   15328: 'Mixinghead 04: Cleaning piston: Front position not reached', class Mixing Head Warning, trigger "Mixinghead_Cpiston4_DBW_40" bit 3
   15329: 'Mixinghead 04: Cleaning piston: Rear position not reached', class Mixing Head Warning, trigger "Mixinghead_Cpiston4_DBW_40" bit 4
   15330: 'Mixinghead 04: Cleaning piston: Home position not reached', class Mixing Head Warning, trigger "Mixinghead_Cpiston4_DBW_40" bit 5
   15331: 'Mixinghead 04: Cleaning piston:', class Mixing Head Warning, trigger "Mixinghead_Cpiston4_DBW_40" bit 6
   15332: 'Mixinghead 04: Cleaning piston:', class Mixing Head Warning, trigger "Mixinghead_Cpiston4_DBW_40" bit 7
   15340: 'Mixinghead 04: Connection 01: Temperature recording: Measuring value outside measuring range', class Mixing Head Warning, trigger "Mixinghead_Temperature_MH4_Con1_DBW76" bit 8
   15341: 'Mixinghead 04: Connection 01: Temperature recording: Warning, value exceeded', class Mixing Head Warning, trigger "Mixinghead_Temperature_MH4_Con1_DBW76" bit 9
   15342: 'Mixinghead 04: Connection 01: Temperature recording: Warning, value undershot', class Mixing Head Warning, trigger "Mixinghead_Temperature_MH4_Con1_DBW76" bit 10
   15343: 'Mixinghead 04: Connection 01: Temperature recording: Fault, value exceeded', class Mixing Head Errors, trigger "Mixinghead_Temperature_MH4_Con1_DBW76" bit 11
   15344: 'Mixinghead 04: Connection 01: Temperature recording: Fault, value undershot', class Mixing Head Errors, trigger "Mixinghead_Temperature_MH4_Con1_DBW76" bit 12
   15345: 'Mixinghead 04: Connection 02: Temperature recording: Measuring value outside measuring range', class Mixing Head Warning, trigger "Mixinghead_Temperature_MH4_Con2_DBW110" bit 8
   15346: 'Mixinghead 04: Connection 02: Temperature recording: Warning, value exceeded', class Mixing Head Warning, trigger "Mixinghead_Temperature_MH4_Con2_DBW110" bit 9
   15347: 'Mixinghead 04: Connection 02: Temperature recording: Warning, value undershot', class Mixing Head Warning, trigger "Mixinghead_Temperature_MH4_Con2_DBW110" bit 10
   15348: 'Mixinghead 04: Connection 02: Temperature recording: Fault, value exceeded', class Mixing Head Errors, trigger "Mixinghead_Temperature_MH4_Con2_DBW110" bit 11
   15349: 'Mixinghead 04: Connection 02: Temperature recording: Fault, value undershot', class Mixing Head Errors, trigger "Mixinghead_Temperature_MH4_Con2_DBW110" bit 12
   15350: 'Mixinghead 04: Connection 03: Temperature recording: Measuring value outside measuring range', class Mixing Head Warning, trigger "Mixinghead_Temperature_MH4_Con3_DBW144" bit 8
   15351: 'Mixinghead 04: Connection 03: Temperature recording: Warning, value exceeded', class Mixing Head Warning, trigger "Mixinghead_Temperature_MH4_Con3_DBW144" bit 9
   15352: 'Mixinghead 04: Connection 03: Temperature recording: Warning, value undershot', class Mixing Head Warning, trigger "Mixinghead_Temperature_MH4_Con3_DBW144" bit 10
   15353: 'Mixinghead 04: Connection 03: Temperature recording: Fault, value exceeded', class Mixing Head Errors, trigger "Mixinghead_Temperature_MH4_Con3_DBW144" bit 11
   15354: 'Mixinghead 04: Connection 03: Temperature recording: Fault, value undershot', class Mixing Head Errors, trigger "Mixinghead_Temperature_MH4_Con3_DBW144" bit 12
   15355: 'Mixinghead 04: Connection 04: Temperature recording: Measuring value outside measuring range', class Mixing Head Warning, trigger "Mixinghead_Temperature_MH4_Con4_DBW178" bit 8
   15356: 'Mixinghead 04: Connection 04: Temperature recording: Warning, value exceeded', class Mixing Head Warning, trigger "Mixinghead_Temperature_MH4_Con4_DBW178" bit 9
   15357: 'Mixinghead 04: Connection 04: Temperature recording: Warning, value undershot', class Mixing Head Warning, trigger "Mixinghead_Temperature_MH4_Con4_DBW178" bit 10
   15358: 'Mixinghead 04: Connection 04: Temperature recording: Fault, value exceeded', class Mixing Head Errors, trigger "Mixinghead_Temperature_MH4_Con4_DBW178" bit 11
   15359: 'Mixinghead 04: Connection 04: Temperature recording: Fault, value undershot', class Mixing Head Errors, trigger "Mixinghead_Temperature_MH4_Con4_DBW178" bit 12
   15360: 'Mixinghead 04: Connection 05: Temperature recording: Measuring value outside measuring range', class Mixing Head Warning, trigger "Mixinghead_Temperature_MH4_Con5_DBW212" bit 8
   15361: 'Mixinghead 04: Connection 05: Temperature recording: Warning, value exceeded', class Mixing Head Warning, trigger "Mixinghead_Temperature_MH4_Con5_DBW212" bit 9
   15362: 'Mixinghead 04: Connection 05: Temperature recording: Warning, value undershot', class Mixing Head Warning, trigger "Mixinghead_Temperature_MH4_Con5_DBW212" bit 10
   15363: 'Mixinghead 04: Connection 05: Temperature recording: Fault, value exceeded', class Mixing Head Errors, trigger "Mixinghead_Temperature_MH4_Con5_DBW212" bit 11
   15364: 'Mixinghead 04: Connection 05: Temperature recording: Fault, value undershot', class Mixing Head Errors, trigger "Mixinghead_Temperature_MH4_Con5_DBW212" bit 12
   15365: 'Mixinghead 04: Connection 06: Temperature recording: Measuring value outside measuring range', class Mixing Head Warning, trigger "Mixinghead_Temperature_MH4_Con6_DBW246" bit 8
   15366: 'Mixinghead 04: Connection 06: Temperature recording: Warning, value exceeded', class Mixing Head Warning, trigger "Mixinghead_Temperature_MH4_Con6_DBW246" bit 9
   15367: 'Mixinghead 04: Connection 06: Temperature recording: Warning, value undershot', class Mixing Head Warning, trigger "Mixinghead_Temperature_MH4_Con6_DBW246" bit 10
   15368: 'Mixinghead 04: Connection 06: Temperature recording: Fault, value exceeded', class Mixing Head Errors, trigger "Mixinghead_Temperature_MH4_Con6_DBW246" bit 11
   15369: 'Mixinghead 04: Connection 06: Temperature recording: Fault, value undershot', class Mixing Head Errors, trigger "Mixinghead_Temperature_MH4_Con6_DBW246" bit 12
   15370: 'Mixinghead 04: Connection 01: Pressure recording: Measuring value outside measuring range', class Mixing Head Warning, trigger "Mixinghead_Pressure_MH4_Con1_DBW280" bit 8
   15371: 'Mixinghead 04: Connection 01: Pressure recording: Warning, value exceeded', class Mixing Head Warning, trigger "Mixinghead_Pressure_MH4_Con1_DBW280" bit 9
   15372: 'Mixinghead 04: Connection 01: Pressure recording: Warning, value undershot', class Mixing Head Warning, trigger "Mixinghead_Pressure_MH4_Con1_DBW280" bit 10
   15373: 'Mixinghead 04: Connection 01: Pressure recording: Fault, value exceeded', class Mixing Head Errors, trigger "Mixinghead_Pressure_MH4_Con1_DBW280" bit 11
   15374: 'Mixinghead 04: Connection 01: Pressure recording: Fault, value undershot', class Mixing Head Errors, trigger "Mixinghead_Pressure_MH4_Con1_DBW280" bit 12
   15375: 'Mixinghead 04: Connection 02: Pressure recording: Measuring value outside measuring range', class Mixing Head Warning, trigger "Mixinghead_Pressure_MH4_Con2_DBW314" bit 8
   15376: 'Mixinghead 04: Connection 02: Pressure recording: Warning, value exceeded', class Mixing Head Warning, trigger "Mixinghead_Pressure_MH4_Con2_DBW314" bit 9
   15377: 'Mixinghead 04: Connection 02: Pressure recording: Warning, value undershot', class Mixing Head Warning, trigger "Mixinghead_Pressure_MH4_Con2_DBW314" bit 10
   15378: 'Mixinghead 04: Connection 02: Pressure recording: Fault, value exceeded', class Mixing Head Errors, trigger "Mixinghead_Pressure_MH4_Con2_DBW314" bit 11
   15379: 'Mixinghead 04: Connection 02: Pressure recording: Fault, value undershot', class Mixing Head Errors, trigger "Mixinghead_Pressure_MH4_Con2_DBW314" bit 12
   15380: 'Mixinghead 04: Connection 03: Pressure recording: Measuring value outside measuring range', class Mixing Head Warning, trigger "Mixinghead_Pressure_MH4_Con3_DBW348" bit 8
   15381: 'Mixinghead 04: Connection 03: Pressure recording: Warning, value exceeded', class Mixing Head Warning, trigger "Mixinghead_Pressure_MH4_Con3_DBW348" bit 9
   15382: 'Mixinghead 04: Connection 03: Pressure recording: Warning, value undershot', class Mixing Head Warning, trigger "Mixinghead_Pressure_MH4_Con3_DBW348" bit 10
   15383: 'Mixinghead 04: Connection 03: Pressure recording: Fault, value exceeded', class Mixing Head Errors, trigger "Mixinghead_Pressure_MH4_Con3_DBW348" bit 11
   15384: 'Mixinghead 04: Connection 03: Pressure recording: Fault, value undershot', class Mixing Head Errors, trigger "Mixinghead_Pressure_MH4_Con3_DBW348" bit 12
   15385: 'Mixinghead 04: Connection 04: Pressure recording: Measuring value outside measuring range', class Mixing Head Warning, trigger "Mixinghead_Pressure_MH4_Con4_DBW382" bit 8
   15386: 'Mixinghead 04: Connection 04: Pressure recording: Warning, value exceeded', class Mixing Head Warning, trigger "Mixinghead_Pressure_MH4_Con4_DBW382" bit 9
   15387: 'Mixinghead 04: Connection 04: Pressure recording: Warning, value undershot', class Mixing Head Warning, trigger "Mixinghead_Pressure_MH4_Con4_DBW382" bit 10
   15388: 'Mixinghead 04: Connection 04: Pressure recording: Fault, value exceeded', class Mixing Head Errors, trigger "Mixinghead_Pressure_MH4_Con4_DBW382" bit 11
   15389: 'Mixinghead 04: Connection 04: Pressure recording: Fault, value undershot', class Mixing Head Errors, trigger "Mixinghead_Pressure_MH4_Con4_DBW382" bit 12
   15390: 'Mixinghead 04: Connection 05: Pressure recording: Measuring value outside measuring range', class Mixing Head Warning, trigger "Mixinghead_Pressure_MH4_Con5_DBW416" bit 8
   15391: 'Mixinghead 04: Connection 05: Pressure recording: Warning, value exceeded', class Mixing Head Warning, trigger "Mixinghead_Pressure_MH4_Con5_DBW416" bit 9
   15392: 'Mixinghead 04: Connection 05: Pressure recording: Warning, value undershot', class Mixing Head Warning, trigger "Mixinghead_Pressure_MH4_Con5_DBW416" bit 10
   15393: 'Mixinghead 04: Connection 05: Pressure recording: Fault, value exceeded', class Mixing Head Errors, trigger "Mixinghead_Pressure_MH4_Con5_DBW416" bit 11
   15394: 'Mixinghead 04: Connection 05: Pressure recording: Fault, value undershot', class Mixing Head Errors, trigger "Mixinghead_Pressure_MH4_Con5_DBW416" bit 12
   15395: 'Mixinghead 04: Connection 06: Pressure recording: Measuring value outside measuring range', class Mixing Head Warning, trigger "Mixinghead_Pressure_MH4_Con6_DBW450" bit 8
   15396: 'Mixinghead 04: Connection 06: Pressure recording: Warning, value exceeded', class Mixing Head Warning, trigger "Mixinghead_Pressure_MH4_Con6_DBW450" bit 9
   15397: 'Mixinghead 04: Connection 06: Pressure recording: Warning, value undershot', class Mixing Head Warning, trigger "Mixinghead_Pressure_MH4_Con6_DBW450" bit 10
   15398: 'Mixinghead 04: Connection 06: Pressure recording: Fault, value exceeded', class Mixing Head Errors, trigger "Mixinghead_Pressure_MH4_Con6_DBW450" bit 11
   15399: 'Mixinghead 04: Connection 06: Pressure recording: Fault, value undershot', class Mixing Head Errors, trigger "Mixinghead_Pressure_MH4_Con6_DBW450" bit 12
   15401: 'Mixinghead 05: Mixinghead does not open', class Mixing Head Errors, trigger "Mixinghead_MHControl5_DBW_10" bit 8
   15402: 'Mixinghead 05: Mixinghead does not close', class Mixing Head Errors, trigger "Mixinghead_MHControl5_DBW_10" bit 9
   15403: 'Mixinghead 05: Entry cancelled', class Mixing Head Warning, trigger "Mixinghead_MHControl5_DBW_10" bit 10
   15404: 'Mixinghead 05: Mixinghead open without activation', class Mixing Head Errors, trigger "Mixinghead_MHControl5_DBW_10" bit 11
   15405: 'Mixinghead 05: Mixinghead close during entry', class Mixing Head Warning, trigger "Mixinghead_MHControl5_DBW_10" bit 12
   15406: 'Mixinghead 05: Warning, shot time too short', class Mixing Head Warning, trigger "Mixinghead_MHControl5_DBW_10" bit 13
   15407: 'Mixinghead 05: Warning , shot time too long', class Mixing Head Warning, trigger "Mixinghead_MHControl5_DBW_10" bit 14
   15408: 'Mixinghead 05: Fault, shot time too short', class Mixing Head Warning, trigger "Mixinghead_MHControl5_DBW_10" bit 15
   15409: 'Mixinghead 05: Mixinghead collides when opening or closing', class Mixing Head Warning, trigger "Mixinghead_MHControl5_DBW_10" bit 0
   15410: 'Mixinghead 05: Runtime monitoring when locking mixing head', class Mixing Head Warning, trigger "Mixinghead_MHControl5_DBW_10" bit 1
   15411: 'Mixinghead 05: Runtime monitoring when unlocking mixing head', class Mixing Head Warning, trigger "Mixinghead_MHControl5_DBW_10" bit 2
   15412: 'Mixinghead 05:', class Mixing Head Warning, trigger "Mixinghead_MHControl5_DBW_10" bit 3
   15413: 'Mixinghead 05:', class Mixing Head Warning, trigger "Mixinghead_MHControl5_DBW_10" bit 4
   15414: 'Mixinghead 05:', class Mixing Head Warning, trigger "Mixinghead_MHControl5_DBW_10" bit 5
   15415: 'Mixinghead 05:', class Mixing Head Warning, trigger "Mixinghead_MHControl5_DBW_10" bit 6
   15416: 'Mixinghead 05: Component required in entry is not enabled at this mixing head', class Mixing Head Errors, trigger "Mixinghead_MHControl5_DBW_10" bit 7
   15417: 'Mixinghead 05: Cleaning piston: Moving out too slow', class Mixing Head Errors, trigger "Mixinghead_Cpiston5_DBW_42" bit 8
   15418: 'Mixinghead 05: Cleaning piston: Moving in too slow', class Mixing Head Errors, trigger "Mixinghead_Cpiston5_DBW_42" bit 9
   15419: 'Mixinghead 05: Cleaning piston: Proximity switch defect', class Mixing Head Errors, trigger "Mixinghead_Cpiston5_DBW_42" bit 10
   15420: 'Mixinghead 05: Cleaning piston: Leaves its home position in entry', class Mixing Head Errors, trigger "Mixinghead_Cpiston5_DBW_42" bit 11
   15421: 'Mixinghead 05: Cleaning piston: Not defined', class Mixing Head Warning, trigger "Mixinghead_Cpiston5_DBW_42" bit 12
   15422: 'Mixinghead 05: Cleaning piston:', class Mixing Head Warning, trigger "Mixinghead_Cpiston5_DBW_42" bit 13
   15423: 'Mixinghead 05: Cleaning piston:', class Mixing Head Warning, trigger "Mixinghead_Cpiston5_DBW_42" bit 14
   15424: 'Mixinghead 05: Cleaning piston:', class Mixing Head Warning, trigger "Mixinghead_Cpiston5_DBW_42" bit 15
   15425: 'Mixinghead 05: Cleaning piston: Controller at upper limit', class Mixing Head Warning, trigger "Mixinghead_Cpiston5_DBW_42" bit 0
   15426: 'Mixinghead 05: Cleaning piston: Controller at lower limit', class Mixing Head Warning, trigger "Mixinghead_Cpiston5_DBW_42" bit 1
   15427: 'Mixinghead 05: Cleaning piston:', class Mixing Head Warning, trigger "Mixinghead_Cpiston5_DBW_42" bit 2
   15428: 'Mixinghead 05: Cleaning piston: Front position not reached', class Mixing Head Warning, trigger "Mixinghead_Cpiston5_DBW_42" bit 3
   15429: 'Mixinghead 05: Cleaning piston: Rear position not reached', class Mixing Head Warning, trigger "Mixinghead_Cpiston5_DBW_42" bit 4
   15430: 'Mixinghead 05: Cleaning piston: Home position not reached', class Mixing Head Warning, trigger "Mixinghead_Cpiston5_DBW_42" bit 5
   15431: 'Mixinghead 05: Cleaning piston:', class Mixing Head Warning, trigger "Mixinghead_Cpiston5_DBW_42" bit 6
   15432: 'Mixinghead 05: Cleaning piston:', class Mixing Head Warning, trigger "Mixinghead_Cpiston5_DBW_42" bit 7
   15440: 'Mixinghead 05: Connection 01: Temperature recording: Measuring value outside measuring range', class Mixing Head Warning, trigger "Mixinghead_Temperature_MH5_Con1_DBW78" bit 8
   15441: 'Mixinghead 05: Connection 01: Temperature recording: Warning, value exceeded', class Mixing Head Warning, trigger "Mixinghead_Temperature_MH5_Con1_DBW78" bit 9
   15442: 'Mixinghead 05: Connection 01: Temperature recording: Warning, value undershot', class Mixing Head Warning, trigger "Mixinghead_Temperature_MH5_Con1_DBW78" bit 10
   15443: 'Mixinghead 05: Connection 01: Temperature recording: Fault, value exceeded', class Mixing Head Errors, trigger "Mixinghead_Temperature_MH5_Con1_DBW78" bit 11
   15444: 'Mixinghead 05: Connection 01: Temperature recording: Fault, value undershot', class Mixing Head Errors, trigger "Mixinghead_Temperature_MH5_Con1_DBW78" bit 12
   15445: 'Mixinghead 05: Connection 02: Temperature recording: Measuring value outside measuring range', class Mixing Head Warning, trigger "Mixinghead_Temperature_MH5_Con2_DBW112" bit 8
   15446: 'Mixinghead 05: Connection 02: Temperature recording: Warning, value exceeded', class Mixing Head Warning, trigger "Mixinghead_Temperature_MH5_Con2_DBW112" bit 9
   15447: 'Mixinghead 05: Connection 02: Temperature recording: Warning, value undershot', class Mixing Head Warning, trigger "Mixinghead_Temperature_MH5_Con2_DBW112" bit 10
   15448: 'Mixinghead 05: Connection 02: Temperature recording: Fault, value exceeded', class Mixing Head Errors, trigger "Mixinghead_Temperature_MH5_Con2_DBW112" bit 11
   15449: 'Mixinghead 05: Connection 02: Temperature recording: Fault, value undershot', class Mixing Head Errors, trigger "Mixinghead_Temperature_MH5_Con2_DBW112" bit 12
   15450: 'Mixinghead 05: Connection 03: Temperature recording: Measuring value outside measuring range', class Mixing Head Warning, trigger "Mixinghead_Temperature_MH5_Con3_DBW146" bit 8
   15451: 'Mixinghead 05: Connection 03: Temperature recording: Warning, value exceeded', class Mixing Head Warning, trigger "Mixinghead_Temperature_MH5_Con3_DBW146" bit 9
   15452: 'Mixinghead 05: Connection 03: Temperature recording: Warning, value undershot', class Mixing Head Warning, trigger "Mixinghead_Temperature_MH5_Con3_DBW146" bit 10
   15453: 'Mixinghead 05: Connection 03: Temperature recording: Fault, value exceeded', class Mixing Head Errors, trigger "Mixinghead_Temperature_MH5_Con3_DBW146" bit 11
   15454: 'Mixinghead 05: Connection 03: Temperature recording: Fault, value undershot', class Mixing Head Errors, trigger "Mixinghead_Temperature_MH5_Con3_DBW146" bit 12
   15455: 'Mixinghead 05: Connection 04: Temperature recording: Measuring value outside measuring range', class Mixing Head Warning, trigger "Mixinghead_Temperature_MH5_Con4_DBW180" bit 8
   15456: 'Mixinghead 05: Connection 04: Temperature recording: Warning, value exceeded', class Mixing Head Warning, trigger "Mixinghead_Temperature_MH5_Con4_DBW180" bit 9
   15457: 'Mixinghead 05: Connection 04: Temperature recording: Warning, value undershot', class Mixing Head Warning, trigger "Mixinghead_Temperature_MH5_Con4_DBW180" bit 10
   15458: 'Mixinghead 05: Connection 04: Temperature recording: Fault, value exceeded', class Mixing Head Errors, trigger "Mixinghead_Temperature_MH5_Con4_DBW180" bit 11
   15459: 'Mixinghead 05: Connection 04: Temperature recording: Fault, value undershot', class Mixing Head Errors, trigger "Mixinghead_Temperature_MH5_Con4_DBW180" bit 12
   15460: 'Mixinghead 05: Connection 05: Temperature recording: Measuring value outside measuring range', class Mixing Head Warning, trigger "Mixinghead_Temperature_MH5_Con5_DBW214" bit 8
   15461: 'Mixinghead 05: Connection 05: Temperature recording: Warning, value exceeded', class Mixing Head Warning, trigger "Mixinghead_Temperature_MH5_Con5_DBW214" bit 9
   15462: 'Mixinghead 05: Connection 05: Temperature recording: Warning, value undershot', class Mixing Head Warning, trigger "Mixinghead_Temperature_MH5_Con5_DBW214" bit 10
   15463: 'Mixinghead 05: Connection 05: Temperature recording: Fault, value exceeded', class Mixing Head Errors, trigger "Mixinghead_Temperature_MH5_Con5_DBW214" bit 11
   15464: 'Mixinghead 05: Connection 05: Temperature recording: Fault, value undershot', class Mixing Head Errors, trigger "Mixinghead_Temperature_MH5_Con5_DBW214" bit 12
   15465: 'Mixinghead 05: Connection 06: Temperature recording: Measuring value outside measuring range', class Mixing Head Warning, trigger "Mixinghead_Temperature_MH5_Con6_DBW248" bit 8
   15466: 'Mixinghead 05: Connection 06: Temperature recording: Warning, value exceeded', class Mixing Head Warning, trigger "Mixinghead_Temperature_MH5_Con6_DBW248" bit 9
   15467: 'Mixinghead 05: Connection 06: Temperature recording: Warning, value undershot', class Mixing Head Warning, trigger "Mixinghead_Temperature_MH5_Con6_DBW248" bit 10
   15468: 'Mixinghead 05: Connection 06: Temperature recording: Fault, value exceeded', class Mixing Head Errors, trigger "Mixinghead_Temperature_MH5_Con6_DBW248" bit 11
   15469: 'Mixinghead 05: Connection 06: Temperature recording: Fault, value undershot', class Mixing Head Errors, trigger "Mixinghead_Temperature_MH5_Con6_DBW248" bit 12
   15470: 'Mixinghead 05: Connection 01: Pressure recording: Measuring value outside measuring range', class Mixing Head Warning, trigger "Mixinghead_Pressure_MH5_Con1_DBW282" bit 8
   15471: 'Mixinghead 05: Connection 01: Pressure recording: Warning, value exceeded', class Mixing Head Warning, trigger "Mixinghead_Pressure_MH5_Con1_DBW282" bit 9
   15472: 'Mixinghead 05: Connection 01: Pressure recording: Warning, value undershot', class Mixing Head Warning, trigger "Mixinghead_Pressure_MH5_Con1_DBW282" bit 10
   15473: 'Mixinghead 05: Connection 01: Pressure recording: Fault, value exceeded', class Mixing Head Errors, trigger "Mixinghead_Pressure_MH5_Con1_DBW282" bit 11
   15474: 'Mixinghead 05: Connection 01: Pressure recording: Fault, value undershot', class Mixing Head Errors, trigger "Mixinghead_Pressure_MH5_Con1_DBW282" bit 12
   15475: 'Mixinghead 05: Connection 02: Pressure recording: Measuring value outside measuring range', class Mixing Head Warning, trigger "Mixinghead_Pressure_MH5_Con2_DBW316" bit 8
   15476: 'Mixinghead 05: Connection 02: Pressure recording: Warning, value exceeded', class Mixing Head Warning, trigger "Mixinghead_Pressure_MH5_Con2_DBW316" bit 9
   15477: 'Mixinghead 05: Connection 02: Pressure recording: Warning, value undershot', class Mixing Head Warning, trigger "Mixinghead_Pressure_MH5_Con2_DBW316" bit 10
   15478: 'Mixinghead 05: Connection 02: Pressure recording: Fault, value exceeded', class Mixing Head Errors, trigger "Mixinghead_Pressure_MH5_Con2_DBW316" bit 11
   15479: 'Mixinghead 05: Connection 02: Pressure recording: Fault, value undershot', class Mixing Head Errors, trigger "Mixinghead_Pressure_MH5_Con2_DBW316" bit 12
   15480: 'Mixinghead 05: Connection 03: Pressure recording: Measuring value outside measuring range', class Mixing Head Warning, trigger "Mixinghead_Pressure_MH5_Con3_DBW350" bit 8
   15481: 'Mixinghead 05: Connection 03: Pressure recording: Warning, value exceeded', class Mixing Head Warning, trigger "Mixinghead_Pressure_MH5_Con3_DBW350" bit 9
   15482: 'Mixinghead 05: Connection 03: Pressure recording: Warning, value undershot', class Mixing Head Warning, trigger "Mixinghead_Pressure_MH5_Con3_DBW350" bit 10
   15483: 'Mixinghead 05: Connection 03: Pressure recording: Fault, value exceeded', class Mixing Head Errors, trigger "Mixinghead_Pressure_MH5_Con3_DBW350" bit 11
   15484: 'Mixinghead 05: Connection 03: Pressure recording: Fault, value undershot', class Mixing Head Errors, trigger "Mixinghead_Pressure_MH5_Con3_DBW350" bit 12
   15485: 'Mixinghead 05: Connection 04: Pressure recording: Measuring value outside measuring range', class Mixing Head Warning, trigger "Mixinghead_Pressure_MH5_Con4_DBW384" bit 8
   15486: 'Mixinghead 05: Connection 04: Pressure recording: Warning, value exceeded', class Mixing Head Warning, trigger "Mixinghead_Pressure_MH5_Con4_DBW384" bit 9
   15487: 'Mixinghead 05: Connection 04: Pressure recording: Warning, value undershot', class Mixing Head Warning, trigger "Mixinghead_Pressure_MH5_Con4_DBW384" bit 10
   15488: 'Mixinghead 05: Connection 04: Pressure recording: Fault, value exceeded', class Mixing Head Errors, trigger "Mixinghead_Pressure_MH5_Con4_DBW384" bit 11
   15489: 'Mixinghead 05: Connection 04: Pressure recording: Fault, value undershot', class Mixing Head Errors, trigger "Mixinghead_Pressure_MH5_Con4_DBW384" bit 12
   15490: 'Mixinghead 05: Connection 05: Pressure recording: Measuring value outside measuring range', class Mixing Head Warning, trigger "Mixinghead_Pressure_MH5_Con5_DBW418" bit 8
   15491: 'Mixinghead 05: Connection 05: Pressure recording: Warning, value exceeded', class Mixing Head Warning, trigger "Mixinghead_Pressure_MH5_Con5_DBW418" bit 9
   15492: 'Mixinghead 05: Connection 05: Pressure recording: Warning, value undershot', class Mixing Head Warning, trigger "Mixinghead_Pressure_MH5_Con5_DBW418" bit 10
   15493: 'Mixinghead 05: Connection 05: Pressure recording: Fault, value exceeded', class Mixing Head Errors, trigger "Mixinghead_Pressure_MH5_Con5_DBW418" bit 11
   15494: 'Mixinghead 05: Connection 05: Pressure recording: Fault, value undershot', class Mixing Head Errors, trigger "Mixinghead_Pressure_MH5_Con5_DBW418" bit 12
   15495: 'Mixinghead 05: Connection 06: Pressure recording: Measuring value outside measuring range', class Mixing Head Warning, trigger "Mixinghead_Pressure_MH5_Con6_DBW452" bit 8
   15496: 'Mixinghead 05: Connection 06: Pressure recording: Warning, value exceeded', class Mixing Head Warning, trigger "Mixinghead_Pressure_MH5_Con6_DBW452" bit 9
   15497: 'Mixinghead 05: Connection 06: Pressure recording: Warning, value undershot', class Mixing Head Warning, trigger "Mixinghead_Pressure_MH5_Con6_DBW452" bit 10
   15498: 'Mixinghead 05: Connection 06: Pressure recording: Fault, value exceeded', class Mixing Head Errors, trigger "Mixinghead_Pressure_MH5_Con6_DBW452" bit 11
   15499: 'Mixinghead 05: Connection 06: Pressure recording: Fault, value undershot', class Mixing Head Errors, trigger "Mixinghead_Pressure_MH5_Con6_DBW452" bit 12
   15501: 'Mixinghead 06: Mixinghead does not open', class Mixing Head Errors, trigger "Mixinghead_MHControl6_DBW_12" bit 8
   15502: 'Mixinghead 06: Mixinghead does not close', class Mixing Head Errors, trigger "Mixinghead_MHControl6_DBW_12" bit 9
   15503: 'Mixinghead 06: Entry cancelled', class Mixing Head Warning, trigger "Mixinghead_MHControl6_DBW_12" bit 10
   15504: 'Mixinghead 06: Mixinghead open without activation', class Mixing Head Errors, trigger "Mixinghead_MHControl6_DBW_12" bit 11
   15505: 'Mixinghead 06: Mixinghead close during entry', class Mixing Head Warning, trigger "Mixinghead_MHControl6_DBW_12" bit 12
   15506: 'Mixinghead 06: Warning, shot time too short', class Mixing Head Warning, trigger "Mixinghead_MHControl6_DBW_12" bit 13
   15507: 'Mixinghead 06: Warning , shot time too long', class Mixing Head Warning, trigger "Mixinghead_MHControl6_DBW_12" bit 14
   15508: 'Mixinghead 06: Fault, shot time too short', class Mixing Head Warning, trigger "Mixinghead_MHControl6_DBW_12" bit 15
   15509: 'Mixinghead 06: Mixinghead collides when opening or closing', class Mixing Head Warning, trigger "Mixinghead_MHControl6_DBW_12" bit 0
   15510: 'Mixinghead 06: Runtime monitoring when locking mixing head', class Mixing Head Warning, trigger "Mixinghead_MHControl6_DBW_12" bit 1
   15511: 'Mixinghead 06: Runtime monitoring when unlocking mixing head', class Mixing Head Warning, trigger "Mixinghead_MHControl6_DBW_12" bit 2
   15512: 'Mixinghead 06:', class Mixing Head Warning, trigger "Mixinghead_MHControl6_DBW_12" bit 3
   15513: 'Mixinghead 06:', class Mixing Head Warning, trigger "Mixinghead_MHControl6_DBW_12" bit 4
   15514: 'Mixinghead 06:', class Mixing Head Warning, trigger "Mixinghead_MHControl6_DBW_12" bit 5
   15515: 'Mixinghead 06:', class Mixing Head Warning, trigger "Mixinghead_MHControl6_DBW_12" bit 6
   15516: 'Mixinghead 06: Component required in entry is not enabled at this mixing head', class Mixing Head Errors, trigger "Mixinghead_MHControl6_DBW_12" bit 7
   15517: 'Mixinghead 06: Cleaning piston: Moving out too slow', class Mixing Head Errors, trigger "Mixinghead_Cpiston6_DBW_44" bit 8
   15518: 'Mixinghead 06: Cleaning piston: Moving in too slow', class Mixing Head Errors, trigger "Mixinghead_Cpiston6_DBW_44" bit 9
   15519: 'Mixinghead 06: Cleaning piston: Proximity switch defect', class Mixing Head Errors, trigger "Mixinghead_Cpiston6_DBW_44" bit 10
   15520: 'Mixinghead 06: Cleaning piston: Leaves its home position in entry', class Mixing Head Errors, trigger "Mixinghead_Cpiston6_DBW_44" bit 11
   15521: 'Mixinghead 06: Cleaning piston: Not defined', class Mixing Head Warning, trigger "Mixinghead_Cpiston6_DBW_44" bit 12
   15522: 'Mixinghead 06: Cleaning piston:', class Mixing Head Warning, trigger "Mixinghead_Cpiston6_DBW_44" bit 13
   15523: 'Mixinghead 06: Cleaning piston:', class Mixing Head Warning, trigger "Mixinghead_Cpiston6_DBW_44" bit 14
   15524: 'Mixinghead 06: Cleaning piston:', class Mixing Head Warning, trigger "Mixinghead_Cpiston6_DBW_44" bit 15
   15525: 'Mixinghead 06: Cleaning piston: Controller at upper limit', class Mixing Head Warning, trigger "Mixinghead_Cpiston6_DBW_44" bit 0
   15526: 'Mixinghead 06: Cleaning piston: Controller at lower limit', class Mixing Head Warning, trigger "Mixinghead_Cpiston6_DBW_44" bit 1
   15527: 'Mixinghead 06: Cleaning piston:', class Mixing Head Warning, trigger "Mixinghead_Cpiston6_DBW_44" bit 2
   15528: 'Mixinghead 06: Cleaning piston: Front position not reached', class Mixing Head Warning, trigger "Mixinghead_Cpiston6_DBW_44" bit 3
   15529: 'Mixinghead 06: Cleaning piston: Rear position not reached', class Mixing Head Warning, trigger "Mixinghead_Cpiston6_DBW_44" bit 4
   15530: 'Mixinghead 06: Cleaning piston: Home position not reached', class Mixing Head Warning, trigger "Mixinghead_Cpiston6_DBW_44" bit 5
   15531: 'Mixinghead 06: Cleaning piston:', class Mixing Head Warning, trigger "Mixinghead_Cpiston6_DBW_44" bit 6
   15532: 'Mixinghead 06: Cleaning piston:', class Mixing Head Warning, trigger "Mixinghead_Cpiston6_DBW_44" bit 7
   15540: 'Mixinghead 06: Connection 01: Temperature recording: Measuring value outside measuring range', class Mixing Head Warning, trigger "Mixinghead_Temperature_MH6_Con1_DBW80" bit 8
   15541: 'Mixinghead 06: Connection 01: Temperature recording: Warning, value exceeded', class Mixing Head Warning, trigger "Mixinghead_Temperature_MH6_Con1_DBW80" bit 9
   15542: 'Mixinghead 06: Connection 01: Temperature recording: Warning, value undershot', class Mixing Head Warning, trigger "Mixinghead_Temperature_MH6_Con1_DBW80" bit 10
   15543: 'Mixinghead 06: Connection 01: Temperature recording: Fault, value exceeded', class Mixing Head Errors, trigger "Mixinghead_Temperature_MH6_Con1_DBW80" bit 11
   15544: 'Mixinghead 06: Connection 01: Temperature recording: Fault, value undershot', class Mixing Head Errors, trigger "Mixinghead_Temperature_MH6_Con1_DBW80" bit 12
   15545: 'Mixinghead 06: Connection 02: Temperature recording: Measuring value outside measuring range', class Mixing Head Warning, trigger "Mixinghead_Temperature_MH6_Con2_DBW114" bit 8
   15546: 'Mixinghead 06: Connection 02: Temperature recording: Warning, value exceeded', class Mixing Head Warning, trigger "Mixinghead_Temperature_MH6_Con2_DBW114" bit 9
   15547: 'Mixinghead 06: Connection 02: Temperature recording: Warning, value undershot', class Mixing Head Warning, trigger "Mixinghead_Temperature_MH6_Con2_DBW114" bit 10
   15548: 'Mixinghead 06: Connection 02: Temperature recording: Fault, value exceeded', class Mixing Head Errors, trigger "Mixinghead_Temperature_MH6_Con2_DBW114" bit 11
   15549: 'Mixinghead 06: Connection 02: Temperature recording: Fault, value undershot', class Mixing Head Errors, trigger "Mixinghead_Temperature_MH6_Con2_DBW114" bit 12
   15550: 'Mixinghead 06: Connection 03: Temperature recording: Measuring value outside measuring range', class Mixing Head Warning, trigger "Mixinghead_Temperature_MH6_Con3_DBW148" bit 8
   15551: 'Mixinghead 06: Connection 03: Temperature recording: Warning, value exceeded', class Mixing Head Warning, trigger "Mixinghead_Temperature_MH6_Con3_DBW148" bit 9
   15552: 'Mixinghead 06: Connection 03: Temperature recording: Warning, value undershot', class Mixing Head Warning, trigger "Mixinghead_Temperature_MH6_Con3_DBW148" bit 10
   15553: 'Mixinghead 06: Connection 03: Temperature recording: Fault, value exceeded', class Mixing Head Errors, trigger "Mixinghead_Temperature_MH6_Con3_DBW148" bit 11
   15554: 'Mixinghead 06: Connection 03: Temperature recording: Fault, value undershot', class Mixing Head Errors, trigger "Mixinghead_Temperature_MH6_Con3_DBW148" bit 12
   15555: 'Mixinghead 06: Connection 04: Temperature recording: Measuring value outside measuring range', class Mixing Head Warning, trigger "Mixinghead_Temperature_MH6_Con4_DBW182" bit 8
   15556: 'Mixinghead 06: Connection 04: Temperature recording: Warning, value exceeded', class Mixing Head Warning, trigger "Mixinghead_Temperature_MH6_Con4_DBW182" bit 9
   15557: 'Mixinghead 06: Connection 04: Temperature recording: Warning, value undershot', class Mixing Head Warning, trigger "Mixinghead_Temperature_MH6_Con4_DBW182" bit 10
   15558: 'Mixinghead 06: Connection 04: Temperature recording: Fault, value exceeded', class Mixing Head Errors, trigger "Mixinghead_Temperature_MH6_Con4_DBW182" bit 11
   15559: 'Mixinghead 06: Connection 04: Temperature recording: Fault, value undershot', class Mixing Head Errors, trigger "Mixinghead_Temperature_MH6_Con4_DBW182" bit 12
   15560: 'Mixinghead 06: Connection 05: Temperature recording: Measuring value outside measuring range', class Mixing Head Warning, trigger "Mixinghead_Temperature_MH6_Con5_DBW216" bit 8
   15561: 'Mixinghead 06: Connection 05: Temperature recording: Warning, value exceeded', class Mixing Head Warning, trigger "Mixinghead_Temperature_MH6_Con5_DBW216" bit 9
   15562: 'Mixinghead 06: Connection 05: Temperature recording: Warning, value undershot', class Mixing Head Warning, trigger "Mixinghead_Temperature_MH6_Con5_DBW216" bit 10
   15563: 'Mixinghead 06: Connection 05: Temperature recording: Fault, value exceeded', class Mixing Head Errors, trigger "Mixinghead_Temperature_MH6_Con5_DBW216" bit 11
   15564: 'Mixinghead 06: Connection 05: Temperature recording: Fault, value undershot', class Mixing Head Errors, trigger "Mixinghead_Temperature_MH6_Con5_DBW216" bit 12
   15565: 'Mixinghead 06: Connection 06: Temperature recording: Measuring value outside measuring range', class Mixing Head Warning, trigger "Mixinghead_Temperature_MH6_Con6_DBW250" bit 8
   15566: 'Mixinghead 06: Connection 06: Temperature recording: Warning, value exceeded', class Mixing Head Warning, trigger "Mixinghead_Temperature_MH6_Con6_DBW250" bit 9
   15567: 'Mixinghead 06: Connection 06: Temperature recording: Warning, value undershot', class Mixing Head Warning, trigger "Mixinghead_Temperature_MH6_Con6_DBW250" bit 10
   15568: 'Mixinghead 06: Connection 06: Temperature recording: Fault, value exceeded', class Mixing Head Errors, trigger "Mixinghead_Temperature_MH6_Con6_DBW250" bit 11
   15569: 'Mixinghead 06: Connection 06: Temperature recording: Fault, value undershot', class Mixing Head Errors, trigger "Mixinghead_Temperature_MH6_Con6_DBW250" bit 12
   15570: 'Mixinghead 06: Connection 01: Pressure recording: Measuring value outside measuring range', class Mixing Head Warning, trigger "Mixinghead_Pressure_MH6_Con1_DBW284" bit 8
   15571: 'Mixinghead 06: Connection 01: Pressure recording: Warning, value exceeded', class Mixing Head Warning, trigger "Mixinghead_Pressure_MH6_Con1_DBW284" bit 9
   15572: 'Mixinghead 06: Connection 01: Pressure recording: Warning, value undershot', class Mixing Head Warning, trigger "Mixinghead_Pressure_MH6_Con1_DBW284" bit 10
   15573: 'Mixinghead 06: Connection 01: Pressure recording: Fault, value exceeded', class Mixing Head Errors, trigger "Mixinghead_Pressure_MH6_Con1_DBW284" bit 11
   15574: 'Mixinghead 06: Connection 01: Pressure recording: Fault, value undershot', class Mixing Head Errors, trigger "Mixinghead_Pressure_MH6_Con1_DBW284" bit 12
   15575: 'Mixinghead 06: Connection 02: Pressure recording: Measuring value outside measuring range', class Mixing Head Warning, trigger "Mixinghead_Pressure_MH6_Con2_DBW318" bit 8
   15576: 'Mixinghead 06: Connection 02: Pressure recording: Warning, value exceeded', class Mixing Head Warning, trigger "Mixinghead_Pressure_MH6_Con2_DBW318" bit 9
   15577: 'Mixinghead 06: Connection 02: Pressure recording: Warning, value undershot', class Mixing Head Warning, trigger "Mixinghead_Pressure_MH6_Con2_DBW318" bit 10
   15578: 'Mixinghead 06: Connection 02: Pressure recording: Fault, value exceeded', class Mixing Head Errors, trigger "Mixinghead_Pressure_MH6_Con2_DBW318" bit 11
   15579: 'Mixinghead 06: Connection 02: Pressure recording: Fault, value undershot', class Mixing Head Errors, trigger "Mixinghead_Pressure_MH6_Con2_DBW318" bit 12
   15580: 'Mixinghead 06: Connection 03: Pressure recording: Measuring value outside measuring range', class Mixing Head Warning, trigger "Mixinghead_Pressure_MH6_Con3_DBW352" bit 8
   15581: 'Mixinghead 06: Connection 03: Pressure recording: Warning, value exceeded', class Mixing Head Warning, trigger "Mixinghead_Pressure_MH6_Con3_DBW352" bit 9
   15582: 'Mixinghead 06: Connection 03: Pressure recording: Warning, value undershot', class Mixing Head Warning, trigger "Mixinghead_Pressure_MH6_Con3_DBW352" bit 10
   15583: 'Mixinghead 06: Connection 03: Pressure recording: Fault, value exceeded', class Mixing Head Errors, trigger "Mixinghead_Pressure_MH6_Con3_DBW352" bit 11
   15584: 'Mixinghead 06: Connection 03: Pressure recording: Fault, value undershot', class Mixing Head Errors, trigger "Mixinghead_Pressure_MH6_Con3_DBW352" bit 12
   15585: 'Mixinghead 06: Connection 04: Pressure recording: Measuring value outside measuring range', class Mixing Head Warning, trigger "Mixinghead_Pressure_MH6_Con4_DBW386" bit 8
   15586: 'Mixinghead 06: Connection 04: Pressure recording: Warning, value exceeded', class Mixing Head Warning, trigger "Mixinghead_Pressure_MH6_Con4_DBW386" bit 9
   15587: 'Mixinghead 06: Connection 04: Pressure recording: Warning, value undershot', class Mixing Head Warning, trigger "Mixinghead_Pressure_MH6_Con4_DBW386" bit 10
   15588: 'Mixinghead 06: Connection 04: Pressure recording: Fault, value exceeded', class Mixing Head Errors, trigger "Mixinghead_Pressure_MH6_Con4_DBW386" bit 11
   15589: 'Mixinghead 06: Connection 04: Pressure recording: Fault, value undershot', class Mixing Head Errors, trigger "Mixinghead_Pressure_MH6_Con4_DBW386" bit 12
   15590: 'Mixinghead 06: Connection 05: Pressure recording: Measuring value outside measuring range', class Mixing Head Warning, trigger "Mixinghead_Pressure_MH6_Con5_DBW420" bit 8
   15591: 'Mixinghead 06: Connection 05: Pressure recording: Warning, value exceeded', class Mixing Head Warning, trigger "Mixinghead_Pressure_MH6_Con5_DBW420" bit 9
   15592: 'Mixinghead 06: Connection 05: Pressure recording: Warning, value undershot', class Mixing Head Warning, trigger "Mixinghead_Pressure_MH6_Con5_DBW420" bit 10
   15593: 'Mixinghead 06: Connection 05: Pressure recording: Fault, value exceeded', class Mixing Head Errors, trigger "Mixinghead_Pressure_MH6_Con5_DBW420" bit 11
   15594: 'Mixinghead 06: Connection 05: Pressure recording: Fault, value undershot', class Mixing Head Errors, trigger "Mixinghead_Pressure_MH6_Con5_DBW420" bit 12
   15595: 'Mixinghead 06: Connection 06: Pressure recording: Measuring value outside measuring range', class Mixing Head Warning, trigger "Mixinghead_Pressure_MH6_Con6_DBW454" bit 8
   15596: 'Mixinghead 06: Connection 06: Pressure recording: Warning, value exceeded', class Mixing Head Warning, trigger "Mixinghead_Pressure_MH6_Con6_DBW454" bit 9
   15597: 'Mixinghead 06: Connection 06: Pressure recording: Warning, value undershot', class Mixing Head Warning, trigger "Mixinghead_Pressure_MH6_Con6_DBW454" bit 10
   15598: 'Mixinghead 06: Connection 06: Pressure recording: Fault, value exceeded', class Mixing Head Errors, trigger "Mixinghead_Pressure_MH6_Con6_DBW454" bit 11
   15599: 'Mixinghead 06: Connection 06: Pressure recording: Fault, value undershot', class Mixing Head Errors, trigger "Mixinghead_Pressure_MH6_Con6_DBW454" bit 12
   15601: 'Mixinghead 07: Mixinghead does not open', class Mixing Head Errors, trigger "Mixinghead_MHControl7_DBW_14" bit 8
   15602: 'Mixinghead 07: Mixinghead does not close', class Mixing Head Errors, trigger "Mixinghead_MHControl7_DBW_14" bit 9
   15603: 'Mixinghead 07: Entry cancelled', class Mixing Head Warning, trigger "Mixinghead_MHControl7_DBW_14" bit 10
   15604: 'Mixinghead 07: Mixinghead open without activation', class Mixing Head Errors, trigger "Mixinghead_MHControl7_DBW_14" bit 11
   15605: 'Mixinghead 07: Mixinghead close during entry', class Mixing Head Warning, trigger "Mixinghead_MHControl7_DBW_14" bit 12
   15606: 'Mixinghead 07: Warning, shot time too short', class Mixing Head Warning, trigger "Mixinghead_MHControl7_DBW_14" bit 13
   15607: 'Mixinghead 07: Warning , shot time too long', class Mixing Head Warning, trigger "Mixinghead_MHControl7_DBW_14" bit 14
   15608: 'Mixinghead 07: Fault, shot time too short', class Mixing Head Warning, trigger "Mixinghead_MHControl7_DBW_14" bit 15
   15609: 'Mixinghead 07: Mixinghead collides when opening or closing', class Mixing Head Warning, trigger "Mixinghead_MHControl7_DBW_14" bit 0
   15610: 'Mixinghead 07: Runtime monitoring when locking mixing head', class Mixing Head Warning, trigger "Mixinghead_MHControl7_DBW_14" bit 1
   15611: 'Mixinghead 07: Runtime monitoring when unlocking mixing head', class Mixing Head Warning, trigger "Mixinghead_MHControl7_DBW_14" bit 2
   15612: 'Mixinghead 07:', class Mixing Head Warning, trigger "Mixinghead_MHControl7_DBW_14" bit 3
   15613: 'Mixinghead 07:', class Mixing Head Warning, trigger "Mixinghead_MHControl7_DBW_14" bit 4
   15614: 'Mixinghead 07:', class Mixing Head Warning, trigger "Mixinghead_MHControl7_DBW_14" bit 5
   15615: 'Mixinghead 07:', class Mixing Head Warning, trigger "Mixinghead_MHControl7_DBW_14" bit 6
   15616: 'Mixinghead 07: Component required in entry is not enabled at this mixing head', class Mixing Head Errors, trigger "Mixinghead_MHControl7_DBW_14" bit 7
   15617: 'Mixinghead 07: Cleaning piston: Moving out too slow', class Mixing Head Errors, trigger "Mixinghead_Cpiston7_DBW_46" bit 8
   15618: 'Mixinghead 07: Cleaning piston: Moving in too slow', class Mixing Head Errors, trigger "Mixinghead_Cpiston7_DBW_46" bit 9
   15619: 'Mixinghead 07: Cleaning piston: Proximity switch defect', class Mixing Head Errors, trigger "Mixinghead_Cpiston7_DBW_46" bit 10
   15620: 'Mixinghead 07: Cleaning piston: Leaves its home position in entry', class Mixing Head Errors, trigger "Mixinghead_Cpiston7_DBW_46" bit 11
   15621: 'Mixinghead 07: Cleaning piston: Not defined', class Mixing Head Warning, trigger "Mixinghead_Cpiston7_DBW_46" bit 12
   15622: 'Mixinghead 07: Cleaning piston:', class Mixing Head Warning, trigger "Mixinghead_Cpiston7_DBW_46" bit 13
   15623: 'Mixinghead 07: Cleaning piston:', class Mixing Head Warning, trigger "Mixinghead_Cpiston7_DBW_46" bit 14
   15624: 'Mixinghead 07: Cleaning piston:', class Mixing Head Warning, trigger "Mixinghead_Cpiston7_DBW_46" bit 15
   15625: 'Mixinghead 07: Cleaning piston: Controller at upper limit', class Mixing Head Warning, trigger "Mixinghead_Cpiston7_DBW_46" bit 0
   15626: 'Mixinghead 07: Cleaning piston: Controller at lower limit', class Mixing Head Warning, trigger "Mixinghead_Cpiston7_DBW_46" bit 1
   15627: 'Mixinghead 07: Cleaning piston:', class Mixing Head Warning, trigger "Mixinghead_Cpiston7_DBW_46" bit 2
   15628: 'Mixinghead 07: Cleaning piston: Front position not reached', class Mixing Head Warning, trigger "Mixinghead_Cpiston7_DBW_46" bit 3
   15629: 'Mixinghead 07: Cleaning piston: Rear position not reached', class Mixing Head Warning, trigger "Mixinghead_Cpiston7_DBW_46" bit 4
   15630: 'Mixinghead 07: Cleaning piston: Home position not reached', class Mixing Head Warning, trigger "Mixinghead_Cpiston7_DBW_46" bit 5
   15631: 'Mixinghead 07: Cleaning piston:', class Mixing Head Warning, trigger "Mixinghead_Cpiston7_DBW_46" bit 6
   15632: 'Mixinghead 07: Cleaning piston:', class Mixing Head Warning, trigger "Mixinghead_Cpiston7_DBW_46" bit 7
   15640: 'Mixinghead 07: Connection 01: Temperature recording: Measuring value outside measuring range', class Mixing Head Warning, trigger "Mixinghead_Temperature_MH7_Con1_DBW82" bit 8
   15641: 'Mixinghead 07: Connection 01: Temperature recording: Warning, value exceeded', class Mixing Head Warning, trigger "Mixinghead_Temperature_MH7_Con1_DBW82" bit 9
   15642: 'Mixinghead 07: Connection 01: Temperature recording: Warning, value undershot', class Mixing Head Warning, trigger "Mixinghead_Temperature_MH7_Con1_DBW82" bit 10
   15643: 'Mixinghead 07: Connection 01: Temperature recording: Fault, value exceeded', class Mixing Head Errors, trigger "Mixinghead_Temperature_MH7_Con1_DBW82" bit 11
   15644: 'Mixinghead 07: Connection 01: Temperature recording: Fault, value undershot', class Mixing Head Errors, trigger "Mixinghead_Temperature_MH7_Con1_DBW82" bit 12
   15645: 'Mixinghead 07: Connection 02: Temperature recording: Measuring value outside measuring range', class Mixing Head Warning, trigger "Mixinghead_Temperature_MH7_Con2_DBW116" bit 8
   15646: 'Mixinghead 07: Connection 02: Temperature recording: Warning, value exceeded', class Mixing Head Warning, trigger "Mixinghead_Temperature_MH7_Con2_DBW116" bit 9
   15647: 'Mixinghead 07: Connection 02: Temperature recording: Warning, value undershot', class Mixing Head Warning, trigger "Mixinghead_Temperature_MH7_Con2_DBW116" bit 10
   15648: 'Mixinghead 07: Connection 02: Temperature recording: Fault, value exceeded', class Mixing Head Errors, trigger "Mixinghead_Temperature_MH7_Con2_DBW116" bit 11
   15649: 'Mixinghead 07: Connection 02: Temperature recording: Fault, value undershot', class Mixing Head Errors, trigger "Mixinghead_Temperature_MH7_Con2_DBW116" bit 12
   15650: 'Mixinghead 07: Connection 03: Temperature recording: Measuring value outside measuring range', class Mixing Head Warning, trigger "Mixinghead_Temperature_MH7_Con3_DBW150" bit 8
   15651: 'Mixinghead 07: Connection 03: Temperature recording: Warning, value exceeded', class Mixing Head Warning, trigger "Mixinghead_Temperature_MH7_Con3_DBW150" bit 9
   15652: 'Mixinghead 07: Connection 03: Temperature recording: Warning, value undershot', class Mixing Head Warning, trigger "Mixinghead_Temperature_MH7_Con3_DBW150" bit 10
   15653: 'Mixinghead 07: Connection 03: Temperature recording: Fault, value exceeded', class Mixing Head Errors, trigger "Mixinghead_Temperature_MH7_Con3_DBW150" bit 11
   15654: 'Mixinghead 07: Connection 03: Temperature recording: Fault, value undershot', class Mixing Head Errors, trigger "Mixinghead_Temperature_MH7_Con3_DBW150" bit 12
   15655: 'Mixinghead 07: Connection 04: Temperature recording: Measuring value outside measuring range', class Mixing Head Warning, trigger "Mixinghead_Temperature_MH7_Con4_DBW184" bit 8
   15656: 'Mixinghead 07: Connection 04: Temperature recording: Warning, value exceeded', class Mixing Head Warning, trigger "Mixinghead_Temperature_MH7_Con4_DBW184" bit 9
   15657: 'Mixinghead 07: Connection 04: Temperature recording: Warning, value undershot', class Mixing Head Warning, trigger "Mixinghead_Temperature_MH7_Con4_DBW184" bit 10
   15658: 'Mixinghead 07: Connection 04: Temperature recording: Fault, value exceeded', class Mixing Head Errors, trigger "Mixinghead_Temperature_MH7_Con4_DBW184" bit 11
   15659: 'Mixinghead 07: Connection 04: Temperature recording: Fault, value undershot', class Mixing Head Errors, trigger "Mixinghead_Temperature_MH7_Con4_DBW184" bit 12
   15660: 'Mixinghead 07: Connection 05: Temperature recording: Measuring value outside measuring range', class Mixing Head Warning, trigger "Mixinghead_Temperature_MH7_Con5_DBW218" bit 8
   15661: 'Mixinghead 07: Connection 05: Temperature recording: Warning, value exceeded', class Mixing Head Warning, trigger "Mixinghead_Temperature_MH7_Con5_DBW218" bit 9
   15662: 'Mixinghead 07: Connection 05: Temperature recording: Warning, value undershot', class Mixing Head Warning, trigger "Mixinghead_Temperature_MH7_Con5_DBW218" bit 10
   15663: 'Mixinghead 07: Connection 05: Temperature recording: Fault, value exceeded', class Mixing Head Errors, trigger "Mixinghead_Temperature_MH7_Con5_DBW218" bit 11
   15664: 'Mixinghead 07: Connection 05: Temperature recording: Fault, value undershot', class Mixing Head Errors, trigger "Mixinghead_Temperature_MH7_Con5_DBW218" bit 12
   15665: 'Mixinghead 07: Connection 06: Temperature recording: Measuring value outside measuring range', class Mixing Head Warning, trigger "Mixinghead_Temperature_MH7_Con6_DBW252" bit 8
   15666: 'Mixinghead 07: Connection 06: Temperature recording: Warning, value exceeded', class Mixing Head Warning, trigger "Mixinghead_Temperature_MH7_Con6_DBW252" bit 9
   15667: 'Mixinghead 07: Connection 06: Temperature recording: Warning, value undershot', class Mixing Head Warning, trigger "Mixinghead_Temperature_MH7_Con6_DBW252" bit 10
   15668: 'Mixinghead 07: Connection 06: Temperature recording: Fault, value exceeded', class Mixing Head Errors, trigger "Mixinghead_Temperature_MH7_Con6_DBW252" bit 11
   15669: 'Mixinghead 07: Connection 06: Temperature recording: Fault, value undershot', class Mixing Head Errors, trigger "Mixinghead_Temperature_MH7_Con6_DBW252" bit 12
   15670: 'Mixinghead 07: Connection 01: Pressure recording: Measuring value outside measuring range', class Mixing Head Warning, trigger "Mixinghead_Pressure_MH7_Con1_DBW286" bit 8
   15671: 'Mixinghead 07: Connection 01: Pressure recording: Warning, value exceeded', class Mixing Head Warning, trigger "Mixinghead_Pressure_MH7_Con1_DBW286" bit 9
   15672: 'Mixinghead 07: Connection 01: Pressure recording: Warning, value undershot', class Mixing Head Warning, trigger "Mixinghead_Pressure_MH7_Con1_DBW286" bit 10
   15673: 'Mixinghead 07: Connection 01: Pressure recording: Fault, value exceeded', class Mixing Head Errors, trigger "Mixinghead_Pressure_MH7_Con1_DBW286" bit 11
   15674: 'Mixinghead 07: Connection 01: Pressure recording: Fault, value undershot', class Mixing Head Errors, trigger "Mixinghead_Pressure_MH7_Con1_DBW286" bit 12
